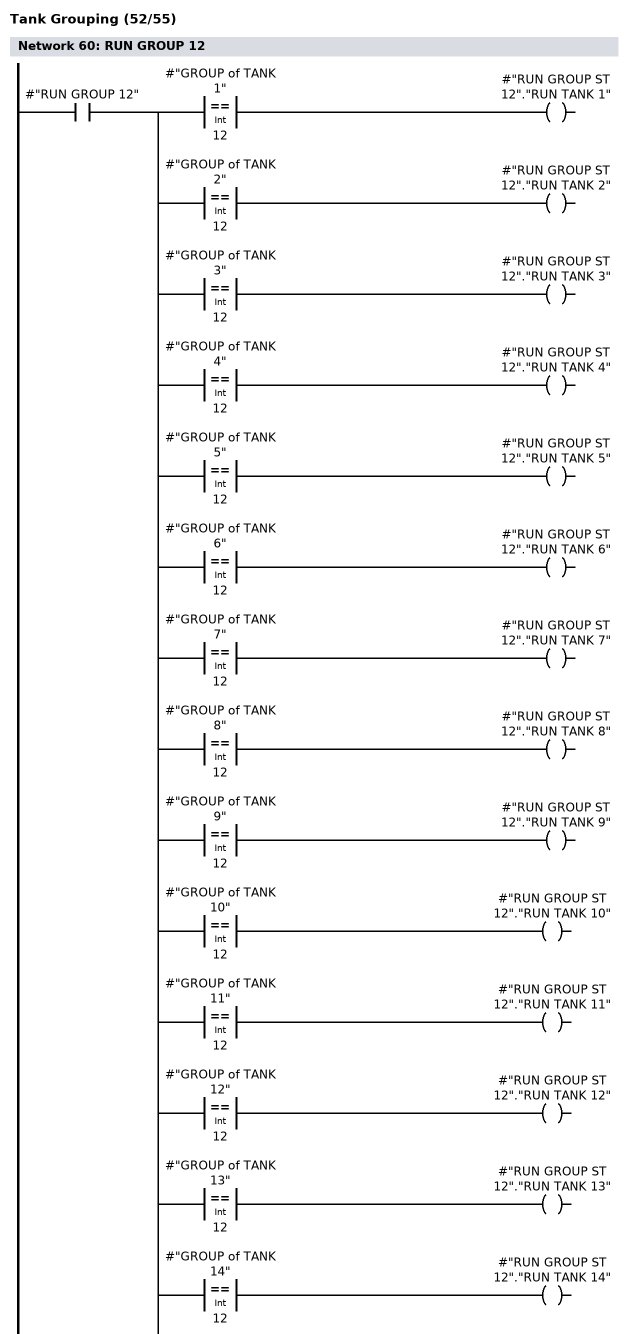
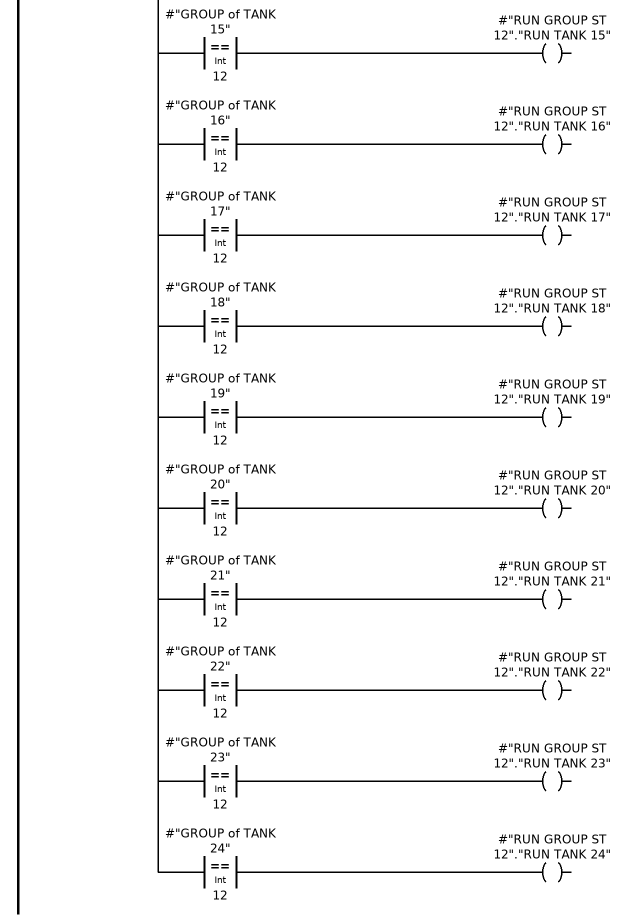
   RUNG wire#powerrail
      Contact( #"RUN GROUP 12" )
      wire#w1
      { S7_Templates := "SrcType := Int" } EQ_Contact(in1 := #"GROUP of TANK 1", in2 := 12)
      Coil( #"RUN GROUP ST 12"."RUN TANK 1" )
   END_RUNG
   RUNG wire#w1
      { S7_Templates := "SrcType := Int" } EQ_Contact(in1 := #"GROUP of TANK 2", in2 := 12)
      Coil( #"RUN GROUP ST 12"."RUN TANK 2" )
   END_RUNG
   RUNG wire#w1
      { S7_Templates := "SrcType := Int" } EQ_Contact(in1 := #"GROUP of TANK 3", in2 := 12)
      Coil( #"RUN GROUP ST 12"."RUN TANK 3" )
   END_RUNG
   RUNG wire#w1
      { S7_Templates := "SrcType := Int" } EQ_Contact(in1 := #"GROUP of TANK 4", in2 := 12)
      Coil( #"RUN GROUP ST 12"."RUN TANK 4" )
   END_RUNG
   RUNG wire#w1
      { S7_Templates := "SrcType := Int" } EQ_Contact(in1 := #"GROUP of TANK 5", in2 := 12)
      Coil( #"RUN GROUP ST 12"."RUN TANK 5" )
   END_RUNG
   RUNG wire#w1
      { S7_Templates := "SrcType := Int" } EQ_Contact(in1 := #"GROUP of TANK 6", in2 := 12)
      Coil( #"RUN GROUP ST 12"."RUN TANK 6" )
   END_RUNG
   RUNG wire#w1
      { S7_Templates := "SrcType := Int" } EQ_Contact(in1 := #"GROUP of TANK 7", in2 := 12)
      Coil( #"RUN GROUP ST 12"."RUN TANK 7" )
   END_RUNG
   RUNG wire#w1
      { S7_Templates := "SrcType := Int" } EQ_Contact(in1 := #"GROUP of TANK 8", in2 := 12)
      Coil( #"RUN GROUP ST 12"."RUN TANK 8" )
   END_RUNG
   RUNG wire#w1
      { S7_Templates := "SrcType := Int" } EQ_Contact(in1 := #"GROUP of TANK 9", in2 := 12)
      Coil( #"RUN GROUP ST 12"."RUN TANK 9" )
   END_RUNG
   RUNG wire#w1
      { S7_Templates := "SrcType := Int" } EQ_Contact(in1 := #"GROUP of TANK 10", in2 := 12)
      Coil( #"RUN GROUP ST 12"."RUN TANK 10" )
   END_RUNG
   RUNG wire#w1
      { S7_Templates := "SrcType := Int" } EQ_Contact(in1 := #"GROUP of TANK 11", in2 := 12)
      Coil( #"RUN GROUP ST 12"."RUN TANK 11" )
   END_RUNG
   RUNG wire#w1
      { S7_Templates := "SrcType := Int" } EQ_Contact(in1 := #"GROUP of TANK 12", in2 := 12)
      Coil( #"RUN GROUP ST 12"."RUN TANK 12" )
   END_RUNG
   RUNG wire#w1
      { S7_Templates := "SrcType := Int" } EQ_Contact(in1 := #"GROUP of TANK 13", in2 := 12)
      Coil( #"RUN GROUP ST 12"."RUN TANK 13" )
   END_RUNG
   RUNG wire#w1
      { S7_Templates := "SrcType := Int" } EQ_Contact(in1 := #"GROUP of TANK 14", in2 := 12)
      Coil( #"RUN GROUP ST 12"."RUN TANK 14" )
   END_RUNG
   RUNG wire#w1
      { S7_Templates := "SrcType := Int" } EQ_Contact(in1 := #"GROUP of TANK 15", in2 := 12)
      Coil( #"RUN GROUP ST 12"."RUN TANK 15" )
   END_RUNG
   RUNG wire#w1
      { S7_Templates := "SrcType := Int" } EQ_Contact(in1 := #"GROUP of TANK 16", in2 := 12)
      Coil( #"RUN GROUP ST 12"."RUN TANK 16" )
   END_RUNG
   RUNG wire#w1
      { S7_Templates := "SrcType := Int" } EQ_Contact(in1 := #"GROUP of TANK 17", in2 := 12)
      Coil( #"RUN GROUP ST 12"."RUN TANK 17" )
   END_RUNG
   RUNG wire#w1
      { S7_Templates := "SrcType := Int" } EQ_Contact(in1 := #"GROUP of TANK 18", in2 := 12)
      Coil( #"RUN GROUP ST 12"."RUN TANK 18" )
   END_RUNG
   RUNG wire#w1
      { S7_Templates := "SrcType := Int" } EQ_Contact(in1 := #"GROUP of TANK 19", in2 := 12)
      Coil( #"RUN GROUP ST 12"."RUN TANK 19" )
   END_RUNG
   RUNG wire#w1
      { S7_Templates := "SrcType := Int" } EQ_Contact(in1 := #"GROUP of TANK 20", in2 := 12)
      Coil( #"RUN GROUP ST 12"."RUN TANK 20" )
   END_RUNG
   RUNG wire#w1
      { S7_Templates := "SrcType := Int" } EQ_Contact(in1 := #"GROUP of TANK 21", in2 := 12)
      Coil( #"RUN GROUP ST 12"."RUN TANK 21" )
   END_RUNG
   RUNG wire#w1
      { S7_Templates := "SrcType := Int" } EQ_Contact(in1 := #"GROUP of TANK 22", in2 := 12)
      Coil( #"RUN GROUP ST 12"."RUN TANK 22" )
   END_RUNG
   RUNG wire#w1
      { S7_Templates := "SrcType := Int" } EQ_Contact(in1 := #"GROUP of TANK 23", in2 := 12)
      Coil( #"RUN GROUP ST 12"."RUN TANK 23" )
   END_RUNG
   RUNG wire#w1
      { S7_Templates := "SrcType := Int" } EQ_Contact(in1 := #"GROUP of TANK 24", in2 := 12)
      Coil( #"RUN GROUP ST 12"."RUN TANK 24" )
   END_RUNG
   // the same network as SCL:
   #"RUN GROUP ST 12"."RUN TANK 1" := #"RUN GROUP 12" AND (#"GROUP of TANK 1" = 12);
   #"RUN GROUP ST 12"."RUN TANK 2" := #"RUN GROUP 12" AND (#"GROUP of TANK 2" = 12);
   #"RUN GROUP ST 12"."RUN TANK 3" := #"RUN GROUP 12" AND (#"GROUP of TANK 3" = 12);
   #"RUN GROUP ST 12"."RUN TANK 4" := #"RUN GROUP 12" AND (#"GROUP of TANK 4" = 12);
   #"RUN GROUP ST 12"."RUN TANK 5" := #"RUN GROUP 12" AND (#"GROUP of TANK 5" = 12);
   #"RUN GROUP ST 12"."RUN TANK 6" := #"RUN GROUP 12" AND (#"GROUP of TANK 6" = 12);
   #"RUN GROUP ST 12"."RUN TANK 7" := #"RUN GROUP 12" AND (#"GROUP of TANK 7" = 12);
   #"RUN GROUP ST 12"."RUN TANK 8" := #"RUN GROUP 12" AND (#"GROUP of TANK 8" = 12);
   #"RUN GROUP ST 12"."RUN TANK 9" := #"RUN GROUP 12" AND (#"GROUP of TANK 9" = 12);
   #"RUN GROUP ST 12"."RUN TANK 10" := #"RUN GROUP 12" AND (#"GROUP of TANK 10" = 12);
   #"RUN GROUP ST 12"."RUN TANK 11" := #"RUN GROUP 12" AND (#"GROUP of TANK 11" = 12);
   #"RUN GROUP ST 12"."RUN TANK 12" := #"RUN GROUP 12" AND (#"GROUP of TANK 12" = 12);
   #"RUN GROUP ST 12"."RUN TANK 13" := #"RUN GROUP 12" AND (#"GROUP of TANK 13" = 12);
   #"RUN GROUP ST 12"."RUN TANK 14" := #"RUN GROUP 12" AND (#"GROUP of TANK 14" = 12);
   #"RUN GROUP ST 12"."RUN TANK 15" := #"RUN GROUP 12" AND (#"GROUP of TANK 15" = 12);
   #"RUN GROUP ST 12"."RUN TANK 16" := #"RUN GROUP 12" AND (#"GROUP of TANK 16" = 12);
   #"RUN GROUP ST 12"."RUN TANK 17" := #"RUN GROUP 12" AND (#"GROUP of TANK 17" = 12);
   #"RUN GROUP ST 12"."RUN TANK 18" := #"RUN GROUP 12" AND (#"GROUP of TANK 18" = 12);
   #"RUN GROUP ST 12"."RUN TANK 19" := #"RUN GROUP 12" AND (#"GROUP of TANK 19" = 12);
   #"RUN GROUP ST 12"."RUN TANK 20" := #"RUN GROUP 12" AND (#"GROUP of TANK 20" = 12);
   #"RUN GROUP ST 12"."RUN TANK 21" := #"RUN GROUP 12" AND (#"GROUP of TANK 21" = 12);
   #"RUN GROUP ST 12"."RUN TANK 22" := #"RUN GROUP 12" AND (#"GROUP of TANK 22" = 12);
   #"RUN GROUP ST 12"."RUN TANK 23" := #"RUN GROUP 12" AND (#"GROUP of TANK 23" = 12);
   #"RUN GROUP ST 12"."RUN TANK 24" := #"RUN GROUP 12" AND (#"GROUP of TANK 24" = 12);
END_REGION

REGION Network 61: RUN GROUP 13
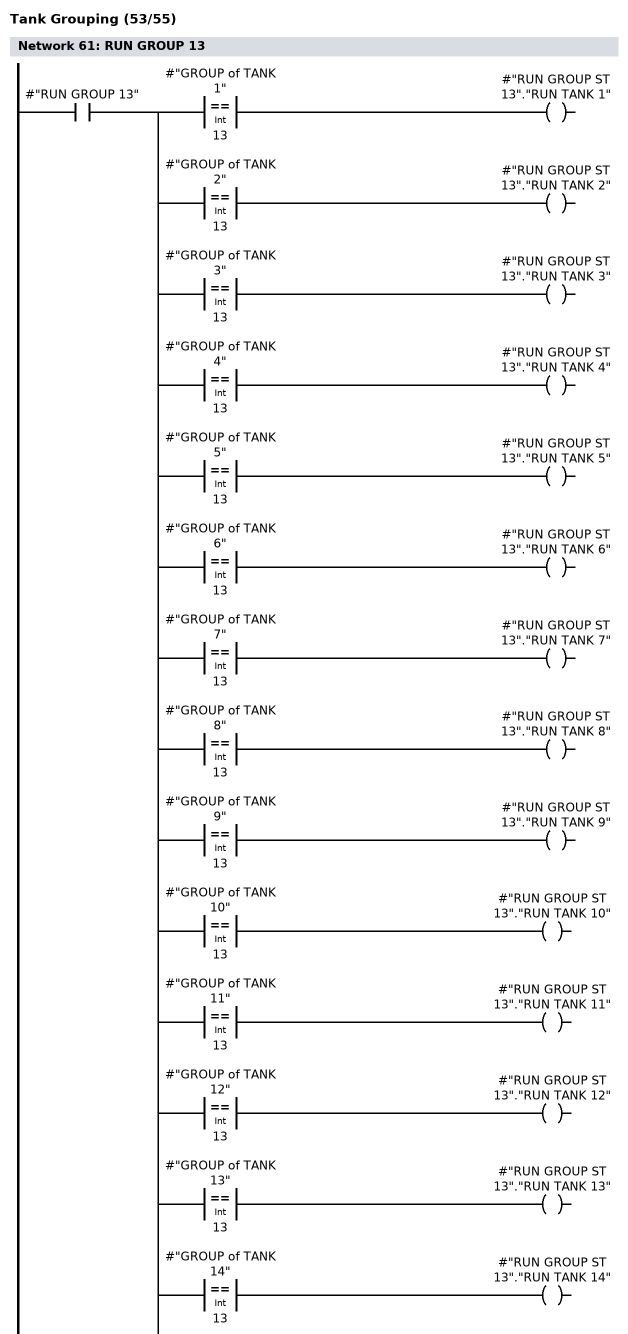
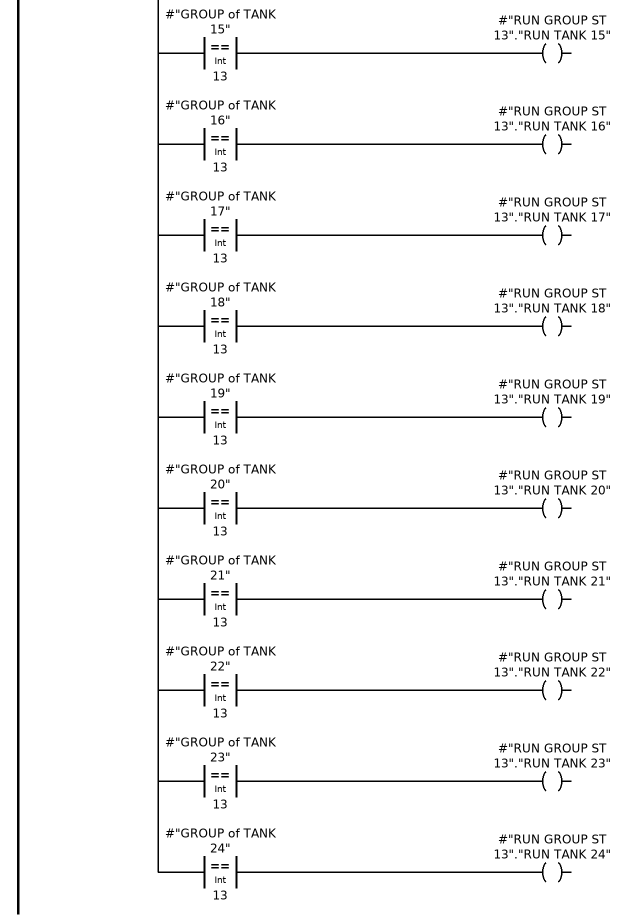
   RUNG wire#powerrail
      Contact( #"RUN GROUP 13" )
      wire#w1
      { S7_Templates := "SrcType := Int" } EQ_Contact(in1 := #"GROUP of TANK 1", in2 := 13)
      Coil( #"RUN GROUP ST 13"."RUN TANK 1" )
   END_RUNG
   RUNG wire#w1
      { S7_Templates := "SrcType := Int" } EQ_Contact(in1 := #"GROUP of TANK 2", in2 := 13)
      Coil( #"RUN GROUP ST 13"."RUN TANK 2" )
   END_RUNG
   RUNG wire#w1
      { S7_Templates := "SrcType := Int" } EQ_Contact(in1 := #"GROUP of TANK 3", in2 := 13)
      Coil( #"RUN GROUP ST 13"."RUN TANK 3" )
   END_RUNG
   RUNG wire#w1
      { S7_Templates := "SrcType := Int" } EQ_Contact(in1 := #"GROUP of TANK 4", in2 := 13)
      Coil( #"RUN GROUP ST 13"."RUN TANK 4" )
   END_RUNG
   RUNG wire#w1
      { S7_Templates := "SrcType := Int" } EQ_Contact(in1 := #"GROUP of TANK 5", in2 := 13)
      Coil( #"RUN GROUP ST 13"."RUN TANK 5" )
   END_RUNG
   RUNG wire#w1
      { S7_Templates := "SrcType := Int" } EQ_Contact(in1 := #"GROUP of TANK 6", in2 := 13)
      Coil( #"RUN GROUP ST 13"."RUN TANK 6" )
   END_RUNG
   RUNG wire#w1
      { S7_Templates := "SrcType := Int" } EQ_Contact(in1 := #"GROUP of TANK 7", in2 := 13)
      Coil( #"RUN GROUP ST 13"."RUN TANK 7" )
   END_RUNG
   RUNG wire#w1
      { S7_Templates := "SrcType := Int" } EQ_Contact(in1 := #"GROUP of TANK 8", in2 := 13)
      Coil( #"RUN GROUP ST 13"."RUN TANK 8" )
   END_RUNG
   RUNG wire#w1
      { S7_Templates := "SrcType := Int" } EQ_Contact(in1 := #"GROUP of TANK 9", in2 := 13)
      Coil( #"RUN GROUP ST 13"."RUN TANK 9" )
   END_RUNG
   RUNG wire#w1
      { S7_Templates := "SrcType := Int" } EQ_Contact(in1 := #"GROUP of TANK 10", in2 := 13)
      Coil( #"RUN GROUP ST 13"."RUN TANK 10" )
   END_RUNG
   RUNG wire#w1
      { S7_Templates := "SrcType := Int" } EQ_Contact(in1 := #"GROUP of TANK 11", in2 := 13)
      Coil( #"RUN GROUP ST 13"."RUN TANK 11" )
   END_RUNG
   RUNG wire#w1
      { S7_Templates := "SrcType := Int" } EQ_Contact(in1 := #"GROUP of TANK 12", in2 := 13)
      Coil( #"RUN GROUP ST 13"."RUN TANK 12" )
   END_RUNG
   RUNG wire#w1
      { S7_Templates := "SrcType := Int" } EQ_Contact(in1 := #"GROUP of TANK 13", in2 := 13)
      Coil( #"RUN GROUP ST 13"."RUN TANK 13" )
   END_RUNG
   RUNG wire#w1
      { S7_Templates := "SrcType := Int" } EQ_Contact(in1 := #"GROUP of TANK 14", in2 := 13)
      Coil( #"RUN GROUP ST 13"."RUN TANK 14" )
   END_RUNG
   RUNG wire#w1
      { S7_Templates := "SrcType := Int" } EQ_Contact(in1 := #"GROUP of TANK 15", in2 := 13)
      Coil( #"RUN GROUP ST 13"."RUN TANK 15" )
   END_RUNG
   RUNG wire#w1
      { S7_Templates := "SrcType := Int" } EQ_Contact(in1 := #"GROUP of TANK 16", in2 := 13)
      Coil( #"RUN GROUP ST 13"."RUN TANK 16" )
   END_RUNG
   RUNG wire#w1
      { S7_Templates := "SrcType := Int" } EQ_Contact(in1 := #"GROUP of TANK 17", in2 := 13)
      Coil( #"RUN GROUP ST 13"."RUN TANK 17" )
   END_RUNG
   RUNG wire#w1
      { S7_Templates := "SrcType := Int" } EQ_Contact(in1 := #"GROUP of TANK 18", in2 := 13)
      Coil( #"RUN GROUP ST 13"."RUN TANK 18" )
   END_RUNG
   RUNG wire#w1
      { S7_Templates := "SrcType := Int" } EQ_Contact(in1 := #"GROUP of TANK 19", in2 := 13)
      Coil( #"RUN GROUP ST 13"."RUN TANK 19" )
   END_RUNG
   RUNG wire#w1
      { S7_Templates := "SrcType := Int" } EQ_Contact(in1 := #"GROUP of TANK 20", in2 := 13)
      Coil( #"RUN GROUP ST 13"."RUN TANK 20" )
   END_RUNG
   RUNG wire#w1
      { S7_Templates := "SrcType := Int" } EQ_Contact(in1 := #"GROUP of TANK 21", in2 := 13)
      Coil( #"RUN GROUP ST 13"."RUN TANK 21" )
   END_RUNG
   RUNG wire#w1
      { S7_Templates := "SrcType := Int" } EQ_Contact(in1 := #"GROUP of TANK 22", in2 := 13)
      Coil( #"RUN GROUP ST 13"."RUN TANK 22" )
   END_RUNG
   RUNG wire#w1
      { S7_Templates := "SrcType := Int" } EQ_Contact(in1 := #"GROUP of TANK 23", in2 := 13)
      Coil( #"RUN GROUP ST 13"."RUN TANK 23" )
   END_RUNG
   RUNG wire#w1
      { S7_Templates := "SrcType := Int" } EQ_Contact(in1 := #"GROUP of TANK 24", in2 := 13)
      Coil( #"RUN GROUP ST 13"."RUN TANK 24" )
   END_RUNG
   // the same network as SCL:
   #"RUN GROUP ST 13"."RUN TANK 1" := #"RUN GROUP 13" AND (#"GROUP of TANK 1" = 13);
   #"RUN GROUP ST 13"."RUN TANK 2" := #"RUN GROUP 13" AND (#"GROUP of TANK 2" = 13);
   #"RUN GROUP ST 13"."RUN TANK 3" := #"RUN GROUP 13" AND (#"GROUP of TANK 3" = 13);
   #"RUN GROUP ST 13"."RUN TANK 4" := #"RUN GROUP 13" AND (#"GROUP of TANK 4" = 13);
   #"RUN GROUP ST 13"."RUN TANK 5" := #"RUN GROUP 13" AND (#"GROUP of TANK 5" = 13);
   #"RUN GROUP ST 13"."RUN TANK 6" := #"RUN GROUP 13" AND (#"GROUP of TANK 6" = 13);
   #"RUN GROUP ST 13"."RUN TANK 7" := #"RUN GROUP 13" AND (#"GROUP of TANK 7" = 13);
   #"RUN GROUP ST 13"."RUN TANK 8" := #"RUN GROUP 13" AND (#"GROUP of TANK 8" = 13);
   #"RUN GROUP ST 13"."RUN TANK 9" := #"RUN GROUP 13" AND (#"GROUP of TANK 9" = 13);
   #"RUN GROUP ST 13"."RUN TANK 10" := #"RUN GROUP 13" AND (#"GROUP of TANK 10" = 13);
   #"RUN GROUP ST 13"."RUN TANK 11" := #"RUN GROUP 13" AND (#"GROUP of TANK 11" = 13);
   #"RUN GROUP ST 13"."RUN TANK 12" := #"RUN GROUP 13" AND (#"GROUP of TANK 12" = 13);
   #"RUN GROUP ST 13"."RUN TANK 13" := #"RUN GROUP 13" AND (#"GROUP of TANK 13" = 13);
   #"RUN GROUP ST 13"."RUN TANK 14" := #"RUN GROUP 13" AND (#"GROUP of TANK 14" = 13);
   #"RUN GROUP ST 13"."RUN TANK 15" := #"RUN GROUP 13" AND (#"GROUP of TANK 15" = 13);
   #"RUN GROUP ST 13"."RUN TANK 16" := #"RUN GROUP 13" AND (#"GROUP of TANK 16" = 13);
   #"RUN GROUP ST 13"."RUN TANK 17" := #"RUN GROUP 13" AND (#"GROUP of TANK 17" = 13);
   #"RUN GROUP ST 13"."RUN TANK 18" := #"RUN GROUP 13" AND (#"GROUP of TANK 18" = 13);
   #"RUN GROUP ST 13"."RUN TANK 19" := #"RUN GROUP 13" AND (#"GROUP of TANK 19" = 13);
   #"RUN GROUP ST 13"."RUN TANK 20" := #"RUN GROUP 13" AND (#"GROUP of TANK 20" = 13);
   #"RUN GROUP ST 13"."RUN TANK 21" := #"RUN GROUP 13" AND (#"GROUP of TANK 21" = 13);
   #"RUN GROUP ST 13"."RUN TANK 22" := #"RUN GROUP 13" AND (#"GROUP of TANK 22" = 13);
   #"RUN GROUP ST 13"."RUN TANK 23" := #"RUN GROUP 13" AND (#"GROUP of TANK 23" = 13);
   #"RUN GROUP ST 13"."RUN TANK 24" := #"RUN GROUP 13" AND (#"GROUP of TANK 24" = 13);
END_REGION

REGION Network 62: RUN GROUP 14
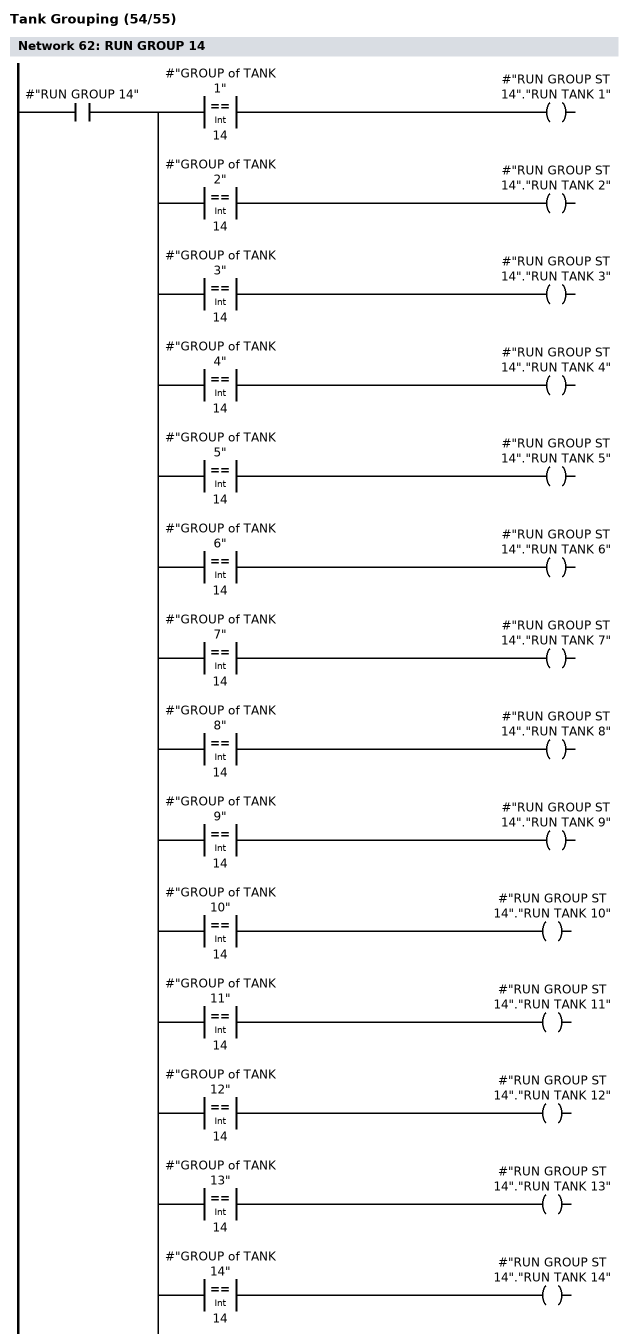
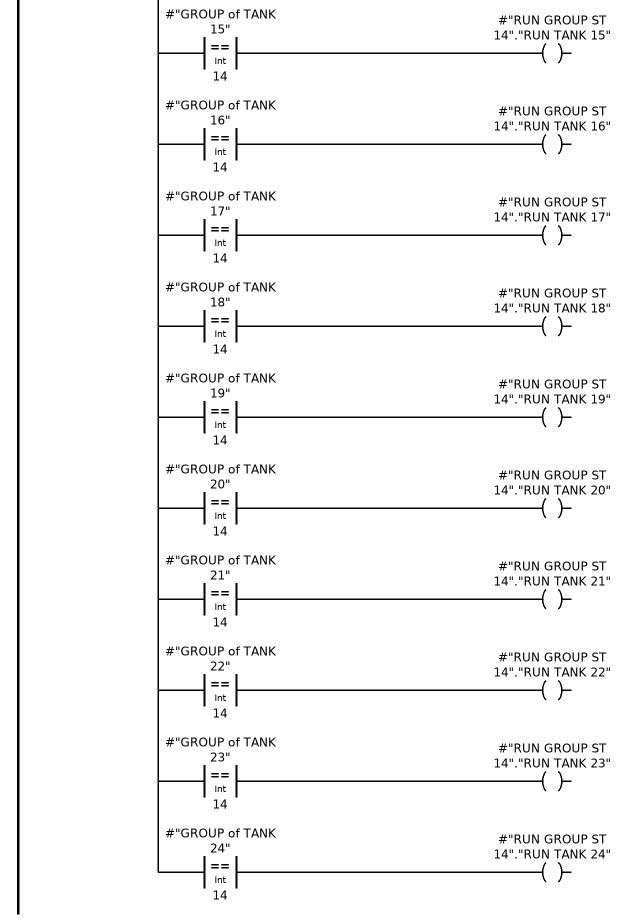
   RUNG wire#powerrail
      Contact( #"RUN GROUP 14" )
      wire#w1
      { S7_Templates := "SrcType := Int" } EQ_Contact(in1 := #"GROUP of TANK 1", in2 := 14)
      Coil( #"RUN GROUP ST 14"."RUN TANK 1" )
   END_RUNG
   RUNG wire#w1
      { S7_Templates := "SrcType := Int" } EQ_Contact(in1 := #"GROUP of TANK 2", in2 := 14)
      Coil( #"RUN GROUP ST 14"."RUN TANK 2" )
   END_RUNG
   RUNG wire#w1
      { S7_Templates := "SrcType := Int" } EQ_Contact(in1 := #"GROUP of TANK 3", in2 := 14)
      Coil( #"RUN GROUP ST 14"."RUN TANK 3" )
   END_RUNG
   RUNG wire#w1
      { S7_Templates := "SrcType := Int" } EQ_Contact(in1 := #"GROUP of TANK 4", in2 := 14)
      Coil( #"RUN GROUP ST 14"."RUN TANK 4" )
   END_RUNG
   RUNG wire#w1
      { S7_Templates := "SrcType := Int" } EQ_Contact(in1 := #"GROUP of TANK 5", in2 := 14)
      Coil( #"RUN GROUP ST 14"."RUN TANK 5" )
   END_RUNG
   RUNG wire#w1
      { S7_Templates := "SrcType := Int" } EQ_Contact(in1 := #"GROUP of TANK 6", in2 := 14)
      Coil( #"RUN GROUP ST 14"."RUN TANK 6" )
   END_RUNG
   RUNG wire#w1
      { S7_Templates := "SrcType := Int" } EQ_Contact(in1 := #"GROUP of TANK 7", in2 := 14)
      Coil( #"RUN GROUP ST 14"."RUN TANK 7" )
   END_RUNG
   RUNG wire#w1
      { S7_Templates := "SrcType := Int" } EQ_Contact(in1 := #"GROUP of TANK 8", in2 := 14)
      Coil( #"RUN GROUP ST 14"."RUN TANK 8" )
   END_RUNG
   RUNG wire#w1
      { S7_Templates := "SrcType := Int" } EQ_Contact(in1 := #"GROUP of TANK 9", in2 := 14)
      Coil( #"RUN GROUP ST 14"."RUN TANK 9" )
   END_RUNG
   RUNG wire#w1
      { S7_Templates := "SrcType := Int" } EQ_Contact(in1 := #"GROUP of TANK 10", in2 := 14)
      Coil( #"RUN GROUP ST 14"."RUN TANK 10" )
   END_RUNG
   RUNG wire#w1
      { S7_Templates := "SrcType := Int" } EQ_Contact(in1 := #"GROUP of TANK 11", in2 := 14)
      Coil( #"RUN GROUP ST 14"."RUN TANK 11" )
   END_RUNG
   RUNG wire#w1
      { S7_Templates := "SrcType := Int" } EQ_Contact(in1 := #"GROUP of TANK 12", in2 := 14)
      Coil( #"RUN GROUP ST 14"."RUN TANK 12" )
   END_RUNG
   RUNG wire#w1
      { S7_Templates := "SrcType := Int" } EQ_Contact(in1 := #"GROUP of TANK 13", in2 := 14)
      Coil( #"RUN GROUP ST 14"."RUN TANK 13" )
   END_RUNG
   RUNG wire#w1
      { S7_Templates := "SrcType := Int" } EQ_Contact(in1 := #"GROUP of TANK 14", in2 := 14)
      Coil( #"RUN GROUP ST 14"."RUN TANK 14" )
   END_RUNG
   RUNG wire#w1
      { S7_Templates := "SrcType := Int" } EQ_Contact(in1 := #"GROUP of TANK 15", in2 := 14)
      Coil( #"RUN GROUP ST 14"."RUN TANK 15" )
   END_RUNG
   RUNG wire#w1
      { S7_Templates := "SrcType := Int" } EQ_Contact(in1 := #"GROUP of TANK 16", in2 := 14)
      Coil( #"RUN GROUP ST 14"."RUN TANK 16" )
   END_RUNG
   RUNG wire#w1
      { S7_Templates := "SrcType := Int" } EQ_Contact(in1 := #"GROUP of TANK 17", in2 := 14)
      Coil( #"RUN GROUP ST 14"."RUN TANK 17" )
   END_RUNG
   RUNG wire#w1
      { S7_Templates := "SrcType := Int" } EQ_Contact(in1 := #"GROUP of TANK 18", in2 := 14)
      Coil( #"RUN GROUP ST 14"."RUN TANK 18" )
   END_RUNG
   RUNG wire#w1
      { S7_Templates := "SrcType := Int" } EQ_Contact(in1 := #"GROUP of TANK 19", in2 := 14)
      Coil( #"RUN GROUP ST 14"."RUN TANK 19" )
   END_RUNG
   RUNG wire#w1
      { S7_Templates := "SrcType := Int" } EQ_Contact(in1 := #"GROUP of TANK 20", in2 := 14)
      Coil( #"RUN GROUP ST 14"."RUN TANK 20" )
   END_RUNG
   RUNG wire#w1
      { S7_Templates := "SrcType := Int" } EQ_Contact(in1 := #"GROUP of TANK 21", in2 := 14)
      Coil( #"RUN GROUP ST 14"."RUN TANK 21" )
   END_RUNG
   RUNG wire#w1
      { S7_Templates := "SrcType := Int" } EQ_Contact(in1 := #"GROUP of TANK 22", in2 := 14)
      Coil( #"RUN GROUP ST 14"."RUN TANK 22" )
   END_RUNG
   RUNG wire#w1
      { S7_Templates := "SrcType := Int" } EQ_Contact(in1 := #"GROUP of TANK 23", in2 := 14)
      Coil( #"RUN GROUP ST 14"."RUN TANK 23" )
   END_RUNG
   RUNG wire#w1
      { S7_Templates := "SrcType := Int" } EQ_Contact(in1 := #"GROUP of TANK 24", in2 := 14)
      Coil( #"RUN GROUP ST 14"."RUN TANK 24" )
   END_RUNG
   // the same network as SCL:
   #"RUN GROUP ST 14"."RUN TANK 1" := #"RUN GROUP 14" AND (#"GROUP of TANK 1" = 14);
   #"RUN GROUP ST 14"."RUN TANK 2" := #"RUN GROUP 14" AND (#"GROUP of TANK 2" = 14);
   #"RUN GROUP ST 14"."RUN TANK 3" := #"RUN GROUP 14" AND (#"GROUP of TANK 3" = 14);
   #"RUN GROUP ST 14"."RUN TANK 4" := #"RUN GROUP 14" AND (#"GROUP of TANK 4" = 14);
   #"RUN GROUP ST 14"."RUN TANK 5" := #"RUN GROUP 14" AND (#"GROUP of TANK 5" = 14);
   #"RUN GROUP ST 14"."RUN TANK 6" := #"RUN GROUP 14" AND (#"GROUP of TANK 6" = 14);
   #"RUN GROUP ST 14"."RUN TANK 7" := #"RUN GROUP 14" AND (#"GROUP of TANK 7" = 14);
   #"RUN GROUP ST 14"."RUN TANK 8" := #"RUN GROUP 14" AND (#"GROUP of TANK 8" = 14);
   #"RUN GROUP ST 14"."RUN TANK 9" := #"RUN GROUP 14" AND (#"GROUP of TANK 9" = 14);
   #"RUN GROUP ST 14"."RUN TANK 10" := #"RUN GROUP 14" AND (#"GROUP of TANK 10" = 14);
   #"RUN GROUP ST 14"."RUN TANK 11" := #"RUN GROUP 14" AND (#"GROUP of TANK 11" = 14);
   #"RUN GROUP ST 14"."RUN TANK 12" := #"RUN GROUP 14" AND (#"GROUP of TANK 12" = 14);
   #"RUN GROUP ST 14"."RUN TANK 13" := #"RUN GROUP 14" AND (#"GROUP of TANK 13" = 14);
   #"RUN GROUP ST 14"."RUN TANK 14" := #"RUN GROUP 14" AND (#"GROUP of TANK 14" = 14);
   #"RUN GROUP ST 14"."RUN TANK 15" := #"RUN GROUP 14" AND (#"GROUP of TANK 15" = 14);
   #"RUN GROUP ST 14"."RUN TANK 16" := #"RUN GROUP 14" AND (#"GROUP of TANK 16" = 14);
   #"RUN GROUP ST 14"."RUN TANK 17" := #"RUN GROUP 14" AND (#"GROUP of TANK 17" = 14);
   #"RUN GROUP ST 14"."RUN TANK 18" := #"RUN GROUP 14" AND (#"GROUP of TANK 18" = 14);
   #"RUN GROUP ST 14"."RUN TANK 19" := #"RUN GROUP 14" AND (#"GROUP of TANK 19" = 14);
   #"RUN GROUP ST 14"."RUN TANK 20" := #"RUN GROUP 14" AND (#"GROUP of TANK 20" = 14);
   #"RUN GROUP ST 14"."RUN TANK 21" := #"RUN GROUP 14" AND (#"GROUP of TANK 21" = 14);
   #"RUN GROUP ST 14"."RUN TANK 22" := #"RUN GROUP 14" AND (#"GROUP of TANK 22" = 14);
   #"RUN GROUP ST 14"."RUN TANK 23" := #"RUN GROUP 14" AND (#"GROUP of TANK 23" = 14);
   #"RUN GROUP ST 14"."RUN TANK 24" := #"RUN GROUP 14" AND (#"GROUP of TANK 24" = 14);
END_REGION

REGION Network 63: Time convertion
   // Last added correction for Offset to be equal with sequence time.
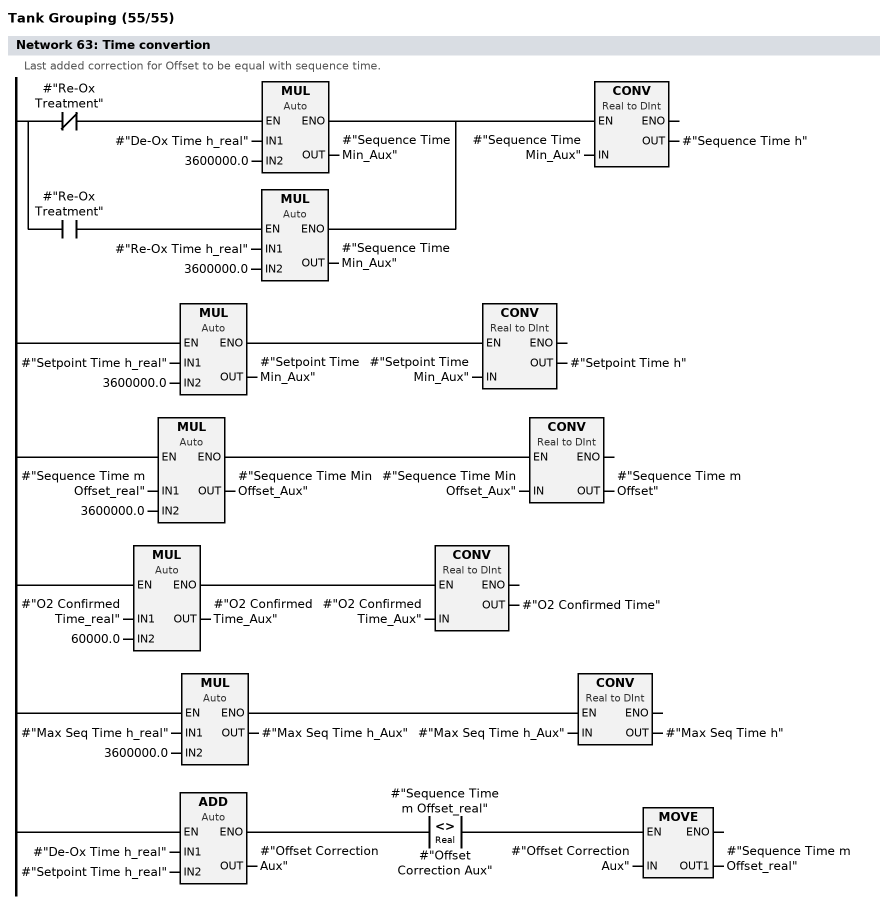
   RUNG wire#powerrail
      I_Contact( #"Re-Ox Treatment" )
      Mul(in1 := #"De-Ox Time h_real", in2 := 3600000.0, out => #"Sequence Time Min_Aux")
      wire#w1
      { S7_Templates := "[SrcType := Real, DestType := DInt]" } Convert(in := #"Sequence Time Min_Aux", out => #"Sequence Time h")
   END_RUNG
   RUNG wire#powerrail
      Contact( #"Re-Ox Treatment" )
      Mul(in1 := #"Re-Ox Time h_real", in2 := 3600000.0, out => #"Sequence Time Min_Aux")
   END_RUNG wire#w1
   RUNG wire#powerrail
      Mul(in1 := #"Setpoint Time h_real", in2 := 3600000.0, out => #"Setpoint Time Min_Aux")
      { S7_Templates := "[SrcType := Real, DestType := DInt]" } Convert(in := #"Setpoint Time Min_Aux", out => #"Setpoint Time h")
   END_RUNG
   RUNG wire#powerrail
      Mul(in1 := #"Sequence Time m Offset_real", in2 := 3600000.0, out => #"Sequence Time Min Offset_Aux")
      { S7_Templates := "[SrcType := Real, DestType := DInt]" } Convert(in := #"Sequence Time Min Offset_Aux", out => #"Sequence Time m Offset")
   END_RUNG
   RUNG wire#powerrail
      Mul(in1 := #"O2 Confirmed Time_real", in2 := 60000.0, out => #"O2 Confirmed Time_Aux")
      { S7_Templates := "[SrcType := Real, DestType := DInt]" } Convert(in := #"O2 Confirmed Time_Aux", out => #"O2 Confirmed Time")
   END_RUNG
   RUNG wire#powerrail
      Mul(in1 := #"Max Seq Time h_real", in2 := 3600000.0, out => #"Max Seq Time h_Aux")
      { S7_Templates := "[SrcType := Real, DestType := DInt]" } Convert(in := #"Max Seq Time h_Aux", out => #"Max Seq Time h")
   END_RUNG
   RUNG wire#powerrail
      Add(in1 := #"De-Ox Time h_real", in2 := #"Setpoint Time h_real", out => #"Offset Correction Aux")
      { S7_Templates := "SrcType := Real" } NE_Contact(in1 := #"Sequence Time m Offset_real", in2 := #"Offset Correction Aux")
      Move(in := #"Offset Correction Aux", out1 => #"Sequence Time m Offset_real")
   END_RUNG
   // the same network as SCL:
   IF NOT #"Re-Ox Treatment" THEN #"Sequence Time Min_Aux" := #"De-Ox Time h_real" * 3600000.0; END_IF;
   IF #"Re-Ox Treatment" THEN #"Sequence Time Min_Aux" := #"Re-Ox Time h_real" * 3600000.0; END_IF;
   IF NOT #"Re-Ox Treatment" OR #"Re-Ox Treatment" THEN
       #"Sequence Time h" := REAL_TO_DINT(#"Sequence Time Min_Aux");
   END_IF;
   #"Setpoint Time Min_Aux" := #"Setpoint Time h_real" * 3600000.0;
   #"Setpoint Time h" := REAL_TO_DINT(#"Setpoint Time Min_Aux");
   #"Sequence Time Min Offset_Aux" := #"Sequence Time m Offset_real" * 3600000.0;
   #"Sequence Time m Offset" := REAL_TO_DINT(#"Sequence Time Min Offset_Aux");
   #"O2 Confirmed Time_Aux" := #"O2 Confirmed Time_real" * 60000.0;
   #"O2 Confirmed Time" := REAL_TO_DINT(#"O2 Confirmed Time_Aux");
   #"Max Seq Time h_Aux" := #"Max Seq Time h_real" * 3600000.0;
   #"Max Seq Time h" := REAL_TO_DINT(#"Max Seq Time h_Aux");
   #"Offset Correction Aux" := #"De-Ox Time h_real" + #"Setpoint Time h_real";
   IF #"Sequence Time m Offset_real" <> #"Offset Correction Aux" THEN
       #"Sequence Time m Offset_real" := #"Offset Correction Aux";
   END_IF;
END_REGION

REGION Network 64: RUN TANK 1
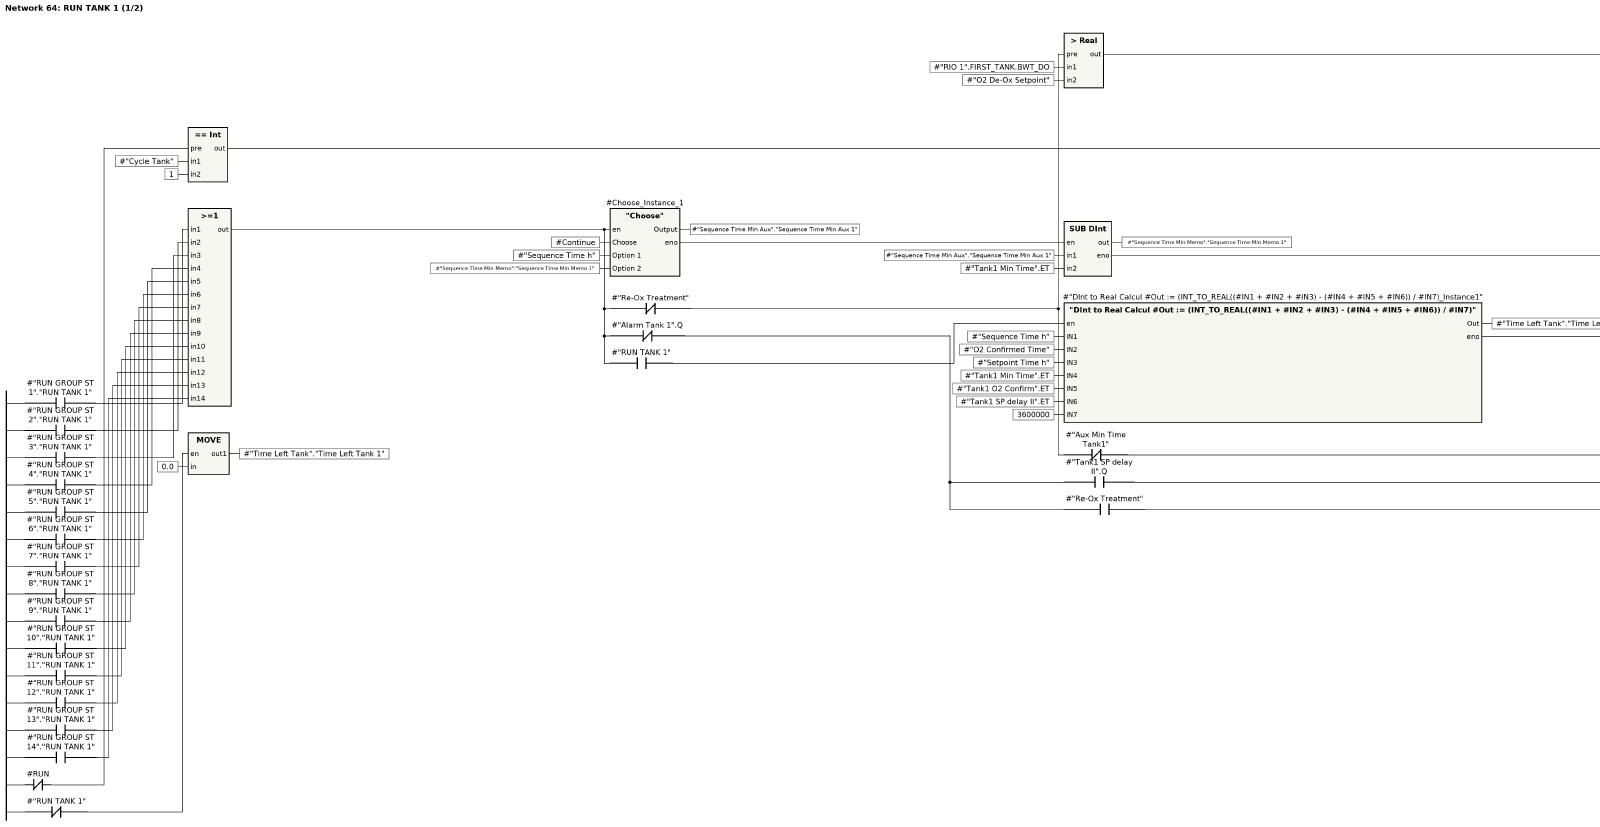
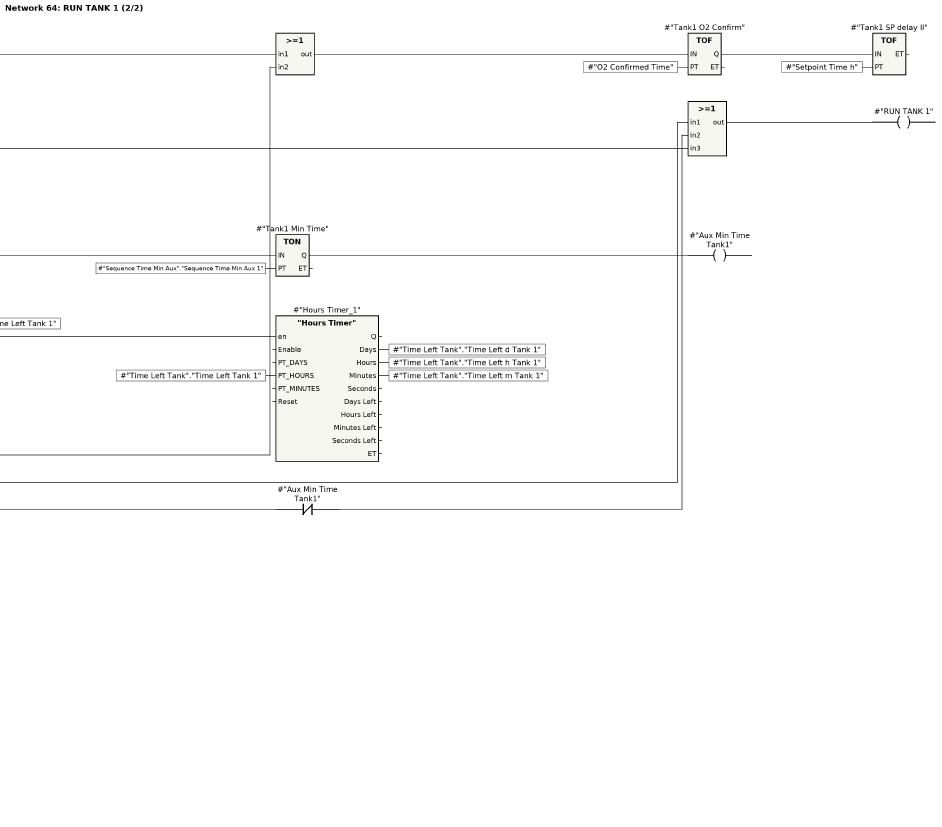
   #_w1 := #"RUN GROUP ST 1"."RUN TANK 1" OR #"RUN GROUP ST 2"."RUN TANK 1" OR #"RUN GROUP ST 3"."RUN TANK 1" OR #"RUN GROUP ST 4"."RUN TANK 1" OR #"RUN GROUP ST 5"."RUN TANK 1" OR #"RUN GROUP ST 6"."RUN TANK 1" OR #"RUN GROUP ST 7"."RUN TANK 1" OR #"RUN GROUP ST 8"."RUN TANK 1" OR #"RUN GROUP ST 9"."RUN TANK 1" OR #"RUN GROUP ST 10"."RUN TANK 1" OR #"RUN GROUP ST 11"."RUN TANK 1" OR #"RUN GROUP ST 12"."RUN TANK 1" OR #"RUN GROUP ST 13"."RUN TANK 1" OR #"RUN GROUP ST 14"."RUN TANK 1";
   #Choose_Instance_1(EN := #_w1,   // "Choose"
                      Choose := #Continue,
                      "Option 1" := #"Sequence Time h",
                      "Option 2" := #"Sequence Time Min Memo"."Sequence Time Min Memo 1",
                      Output => #"Sequence Time Min Aux"."Sequence Time Min Aux 1",
                      ENO => #_w2);
   IF #_w2 THEN
       #"Sequence Time Min Memo"."Sequence Time Min Memo 1" := #"Sequence Time Min Aux"."Sequence Time Min Aux 1" - #"Tank1 Min Time".ET;   // Memory of remained time for use to continue
   END_IF;
   #"Tank1 Min Time"(IN := #_w2, PT := #"Sequence Time Min Aux"."Sequence Time Min Aux 1");   // TON
   #"Aux Min Time Tank1" := #"Tank1 Min Time".Q;
   #"Tank1 O2 Confirm"(IN := #_w1 AND NOT #"Re-Ox Treatment" AND ((#"RIO 1".FIRST_TANK.BWT_DO > #"O2 De-Ox Setpoint") OR NOT #"Aux Min Time Tank1"),   // TOF
                       PT := #"O2 Confirmed Time");
   #"Tank1 SP delay II"(IN := #"Tank1 O2 Confirm".Q, PT := #"Setpoint Time h");   // TOF
   #"DInt to Real Calcul #Out := (INT_TO_REAL((#IN1 + #IN2 + #IN3) - (#IN4 + #IN5 + #IN6)) / #IN7)_Instance1"(EN := #_w1 AND #"RUN TANK 1",   // "DInt to Real Calcul #Out := (INT_TO_REAL((#IN1 + #IN2 + #IN3) - (#IN4 + #IN5 + #IN6)) / #IN7)"
                           IN1 := #"Sequence Time h",
                           IN2 := #"O2 Confirmed Time",
                           IN3 := #"Setpoint Time h",
                           IN4 := #"Tank1 Min Time".ET,
                           IN5 := #"Tank1 O2 Confirm".ET,
                           IN6 := #"Tank1 SP delay II".ET,
                           IN7 := 3600000,
                           Out => #"Time Left Tank"."Time Left Tank 1",
                           ENO => #_w3);
   IF #_w3 THEN
       #"Hours Timer_1"(PT_HOURS := #"Time Left Tank"."Time Left Tank 1",   // "Hours Timer"
                        Days => #"Time Left Tank"."Time Left d Tank 1",
                        Hours => #"Time Left Tank"."Time Left h Tank 1",
                        Minutes => #"Time Left Tank"."Time Left m Tank 1");
   END_IF;
   #"RUN TANK 1" := (#_w1 AND NOT #"Alarm Tank 1".Q AND (#"Tank1 SP delay II".Q OR (#"Re-Ox Treatment" AND NOT #"Aux Min Time Tank1"))) OR (NOT #RUN AND (#"Cycle Tank" = 1));
   IF NOT #"RUN TANK 1" THEN #"Time Left Tank"."Time Left Tank 1" := 0.0; END_IF;
END_REGION

REGION Network 65: RUN TANK 2
